(* Logix 5000 project; controller PLC_MCC1201_220AP1 vendor 1 type 14 code 164 rev 35.11; software revision 35.00; part 12 of 25 *)
(* tags used below, declared in another part *)
   B180 : DINT[10];
   BT181_009 : MESSAGE;
   BT181_010 : MESSAGE;
   C183 : COUNTER[3];
   N124 : DINT[414];
   N125 : DINT[414];
   N126 : DINT[103];
   N127 : DINT[997];
   N128 : DINT[997];
   N177_0 : ALIAS FOR N177[0];
   N184 : DINT[50];
   N184_1 : ALIAS FOR N184[1];
   N184_11 : ALIAS FOR N184[11];
   N184_12 : ALIAS FOR N184[12];
   N184_14 : ALIAS FOR N184[14];
   N184_16 : ALIAS FOR N184[16];
   N184_2 : ALIAS FOR N184[2];
   N184_21 : ALIAS FOR N184[21];
   N184_22 : ALIAS FOR N184[22];
   N184_24 : ALIAS FOR N184[24];
   N184_25 : ALIAS FOR N184[25];
   N184_26 : ALIAS FOR N184[26];
   N184_31 : ALIAS FOR N184[31];
   N184_32 : ALIAS FOR N184[32];
   N184_34 : ALIAS FOR N184[34];
   N184_36 : ALIAS FOR N184[36];
   N184_4 : ALIAS FOR N184[4];
   N184_5 : ALIAS FOR N184[5];
   N184_6 : ALIAS FOR N184[6];
   N26 : DINT[1000];
   T182 : TIMER[11];
   TMP_xAlwaysOFF : BOOL;
(* MainProgram, continued *)

ROUTINE _103_LADDER   (* ladder *)
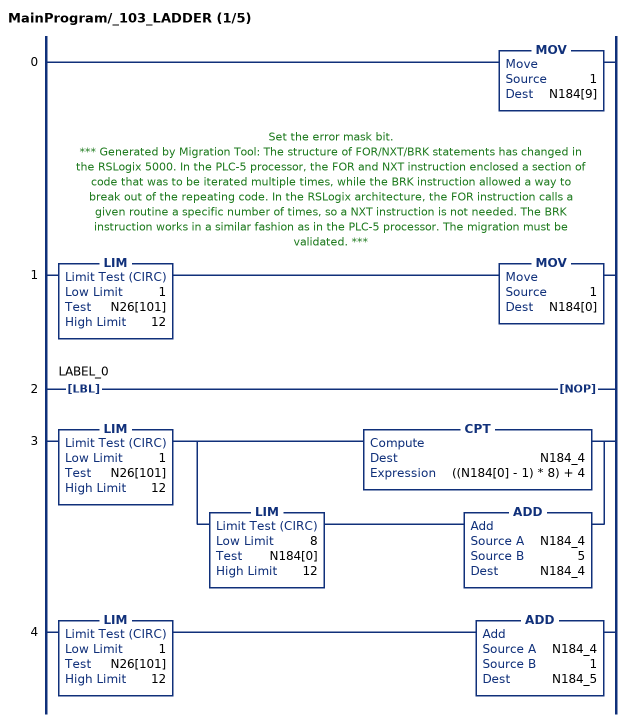
   0: MOV(1,N184[9]);
   // Set the error mask bit.
   // *** Generated by Migration Tool: The structure of FOR/NXT/BRK statements has changed in the RSLogix 5000. In the PLC-5 processor, the FOR and NXT instruction enclosed a section of code that was to be iterated multiple times, while the BRK instruction allowed a way to break out of the repeating code. In the RSLogix architecture, the FOR instruction calls a given routine a specific number of times, so a NXT instruction is not needed. The BRK instruction works in a similar fashion as in the PLC-5 processor. The migration must be validated. ***
   1: LIM(1,N26[101],12)MOV(1,N184[0]);
   2: LBL(LABEL_0)NOP();
   3: LIM(1,N26[101],12)[CPT(N184_4,((N184[0] - 1) * 8) + 4) ,LIM(8,N184[0],12) ADD(N184_4,5,N184_4) ];
   4: LIM(1,N26[101],12)ADD(N184_4,1,N184_5);
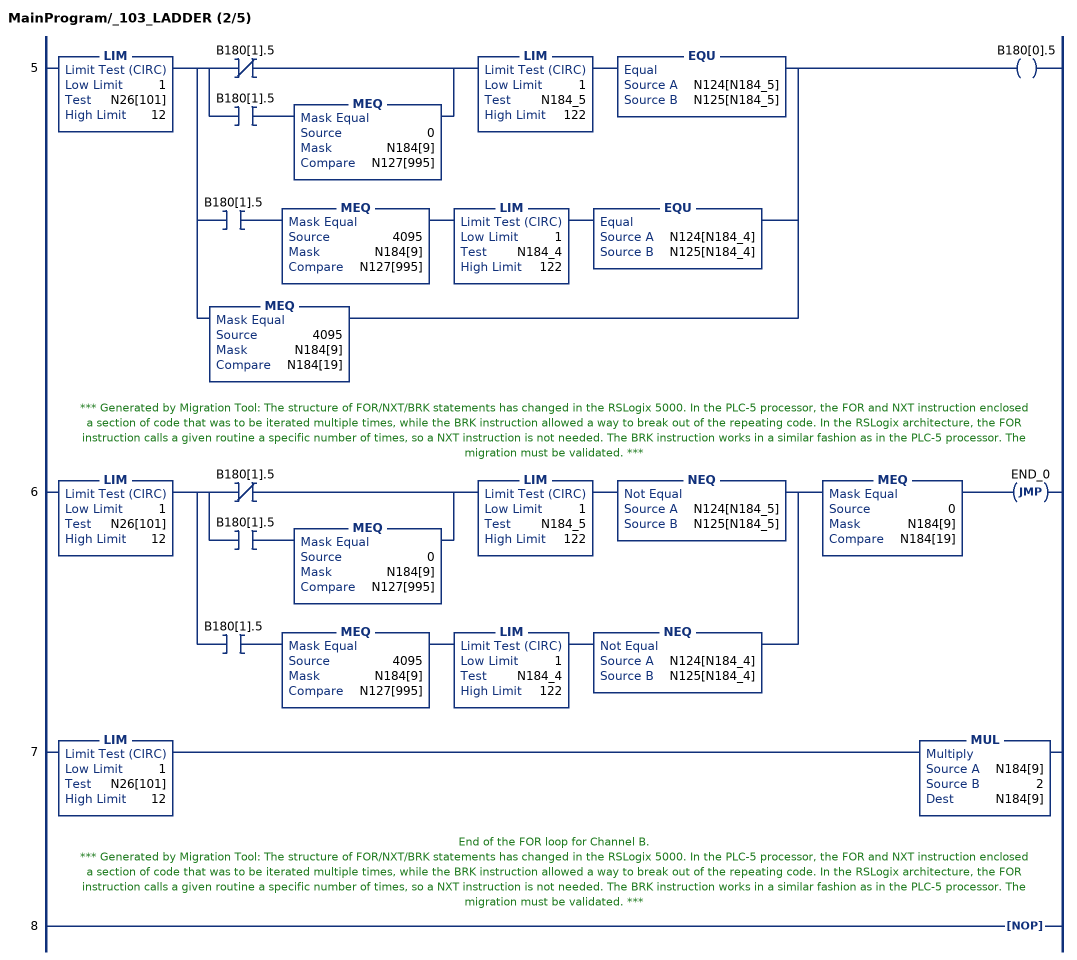
   5: LIM(1,N26[101],12)[[XIO(B180[1].5) ,XIC(B180[1].5) MEQ(0,N184[9],N127[995]) ] LIM(1,N184_5,122) EQU(N124[N184_5],N125[N184_5]) ,XIC(B180[1].5) MEQ(4095,N184[9],N127[995]) LIM(1,N184_4,122) EQU(N124[N184_4],N125[N184_4]) ,MEQ(4095,N184[9],N184[19]) ]OTE(B180[0].5);
   // *** Generated by Migration Tool: The structure of FOR/NXT/BRK statements has changed in the RSLogix 5000. In the PLC-5 processor, the FOR and NXT instruction enclosed a section of code that was to be iterated multiple times, while the BRK instruction allowed a way to break out of the repeating code. In the RSLogix architecture, the FOR instruction calls a given routine a specific number of times, so a NXT instruction is not needed. The BRK instruction works in a similar fashion as in the PLC-5 processor. The migration must be validated. ***
   6: LIM(1,N26[101],12)[[XIO(B180[1].5) ,XIC(B180[1].5) MEQ(0,N184[9],N127[995]) ] LIM(1,N184_5,122) NEQ(N124[N184_5],N125[N184_5]) ,XIC(B180[1].5) MEQ(4095,N184[9],N127[995]) LIM(1,N184_4,122) NEQ(N124[N184_4],N125[N184_4]) ]MEQ(0,N184[9],N184[19])JMP(END_0);
   7: LIM(1,N26[101],12)MUL(N184[9],2,N184[9]);
   // End of the FOR loop for Channel B.
   // *** Generated by Migration Tool: The structure of FOR/NXT/BRK statements has changed in the RSLogix 5000. In the PLC-5 processor, the FOR and NXT instruction enclosed a section of code that was to be iterated multiple times, while the BRK instruction allowed a way to break out of the repeating code. In the RSLogix architecture, the FOR instruction calls a given routine a specific number of times, so a NXT instruction is not needed. The BRK instruction works in a similar fashion as in the PLC-5 processor. The migration must be validated. ***
   8: NOP();
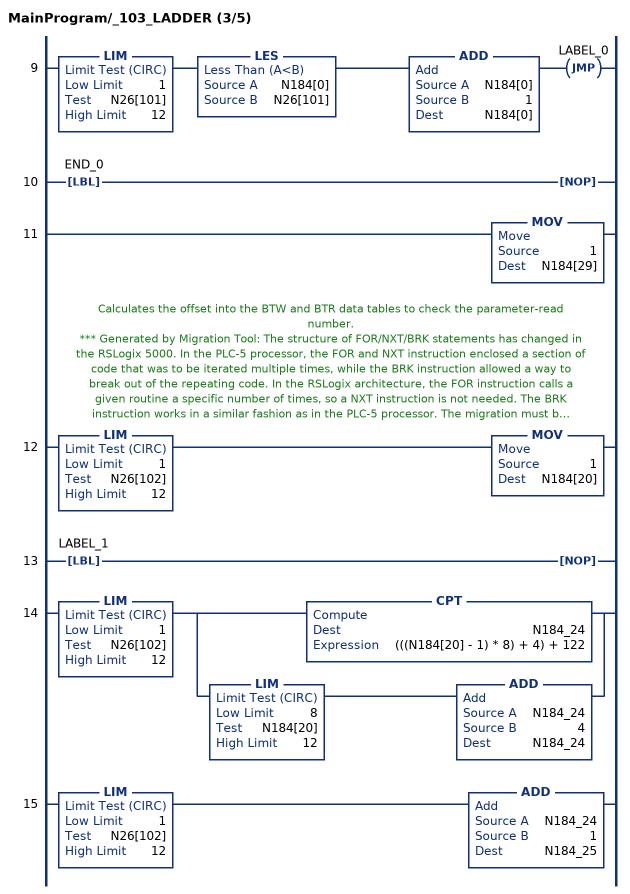
   9: LIM(1,N26[101],12)LES(N184[0],N26[101])ADD(N184[0],1,N184[0])JMP(LABEL_0);
   10: LBL(END_0)NOP();
   11: MOV(1,N184[29]);
   // Calculates the offset into the BTW and BTR data tables to check the parameter-read number.
   // *** Generated by Migration Tool: The structure of FOR/NXT/BRK statements has changed in the RSLogix 5000. In the PLC-5 processor, the FOR and NXT instruction enclosed a section of code that was to be iterated multiple times, while the BRK instruction allowed a way to break out of the repeating code. In the RSLogix architecture, the FOR instruction calls a given routine a specific number of times, so a NXT instruction is not needed. The BRK instruction works in a similar fashion as in the PLC-5 processor. The migration must be validated. ***
   12: LIM(1,N26[102],12)MOV(1,N184[20]);
   13: LBL(LABEL_1)NOP();
   14: LIM(1,N26[102],12)[CPT(N184_24,(((N184[20] - 1) * 8) + 4) + 122) ,LIM(8,N184[20],12) ADD(N184_24,4,N184_24) ];
   15: LIM(1,N26[102],12)ADD(N184_24,1,N184_25);
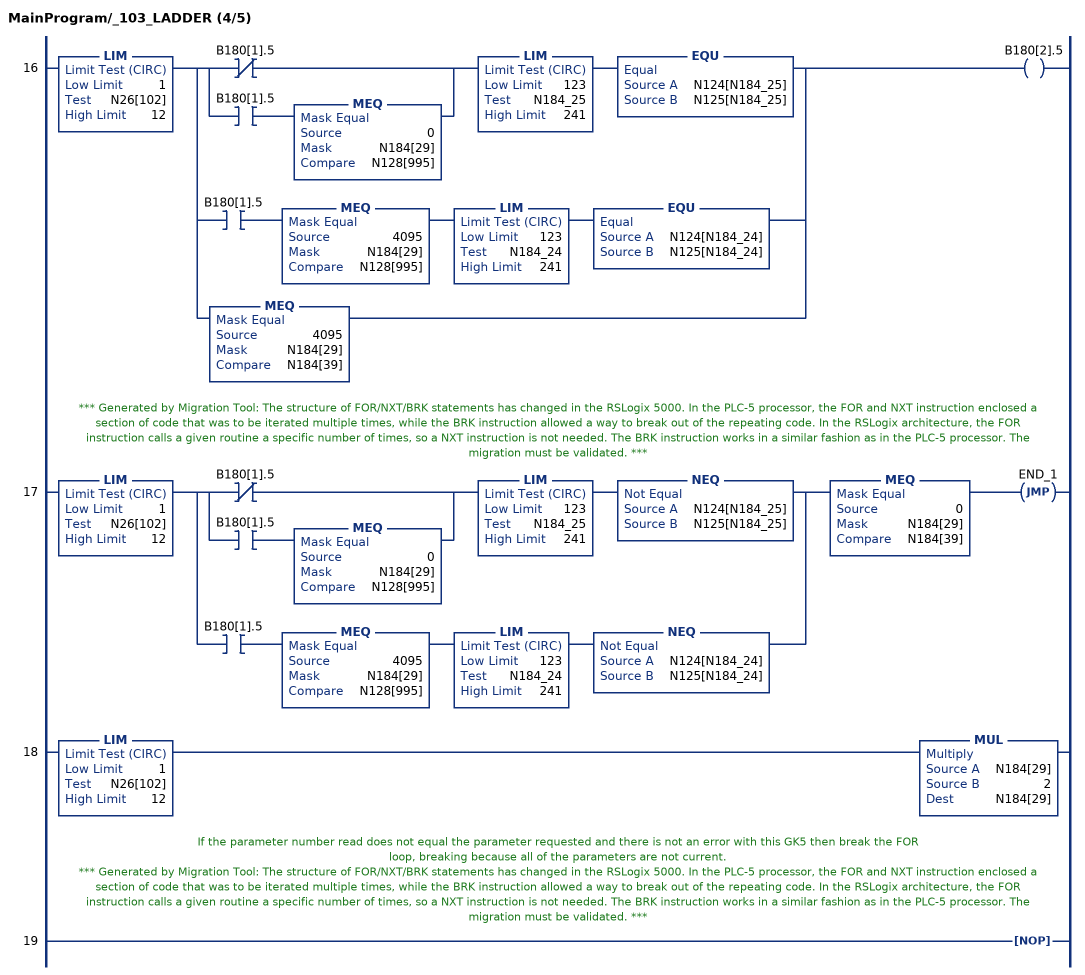
   16: LIM(1,N26[102],12)[[XIO(B180[1].5) ,XIC(B180[1].5) MEQ(0,N184[29],N128[995]) ] LIM(123,N184_25,241) EQU(N124[N184_25],N125[N184_25]) ,XIC(B180[1].5) MEQ(4095,N184[29],N128[995]) LIM(123,N184_24,241) EQU(N124[N184_24],N125[N184_24]) ,MEQ(4095,N184[29],N184[39]) ]OTE(B180[2].5);
   // *** Generated by Migration Tool: The structure of FOR/NXT/BRK statements has changed in the RSLogix 5000. In the PLC-5 processor, the FOR and NXT instruction enclosed a section of code that was to be iterated multiple times, while the BRK instruction allowed a way to break out of the repeating code. In the RSLogix architecture, the FOR instruction calls a given routine a specific number of times, so a NXT instruction is not needed. The BRK instruction works in a similar fashion as in the PLC-5 processor. The migration must be validated. ***
   17: LIM(1,N26[102],12)[[XIO(B180[1].5) ,XIC(B180[1].5) MEQ(0,N184[29],N128[995]) ] LIM(123,N184_25,241) NEQ(N124[N184_25],N125[N184_25]) ,XIC(B180[1].5) MEQ(4095,N184[29],N128[995]) LIM(123,N184_24,241) NEQ(N124[N184_24],N125[N184_24]) ]MEQ(0,N184[29],N184[39])JMP(END_1);
   18: LIM(1,N26[102],12)MUL(N184[29],2,N184[29]);
   // If the parameter number read does not equal the parameter requested and there is not an error with this GK5 then break the FOR
   // loop, breaking because all of the parameters are not current.
   // *** Generated by Migration Tool: The structure of FOR/NXT/BRK statements has changed in the RSLogix 5000. In the PLC-5 processor, the FOR and NXT instruction enclosed a section of code that was to be iterated multiple times, while the BRK instruction allowed a way to break out of the repeating code. In the RSLogix architecture, the FOR instruction calls a given routine a specific number of times, so a NXT instruction is not needed. The BRK instruction works in a similar fashion as in the PLC-5 processor. The migration must be validated. ***
   19: NOP();
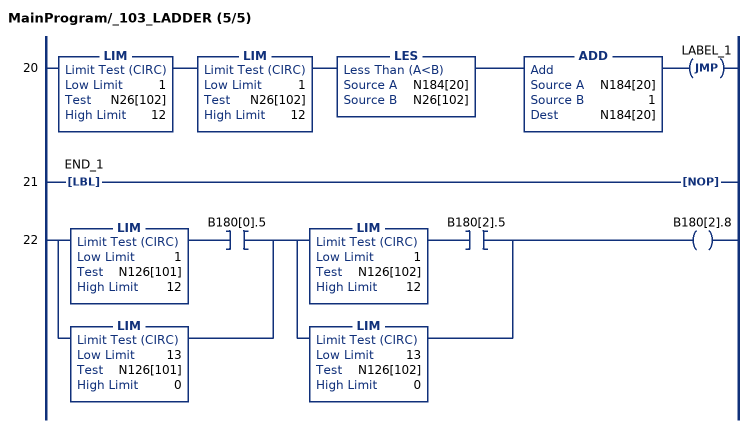
   20: LIM(1,N26[102],12)LIM(1,N26[102],12)LES(N184[20],N26[102])ADD(N184[20],1,N184[20])JMP(LABEL_1);
   21: LBL(END_1)NOP();
   22: [LIM(1,N126[101],12) XIC(B180[0].5) ,LIM(13,N126[101],0) ][LIM(1,N126[102],12) XIC(B180[2].5) ,LIM(13,N126[102],0) ]OTE(B180[2].8);
END_ROUTINE

ROUTINE _104_LADDER   (* ladder *)
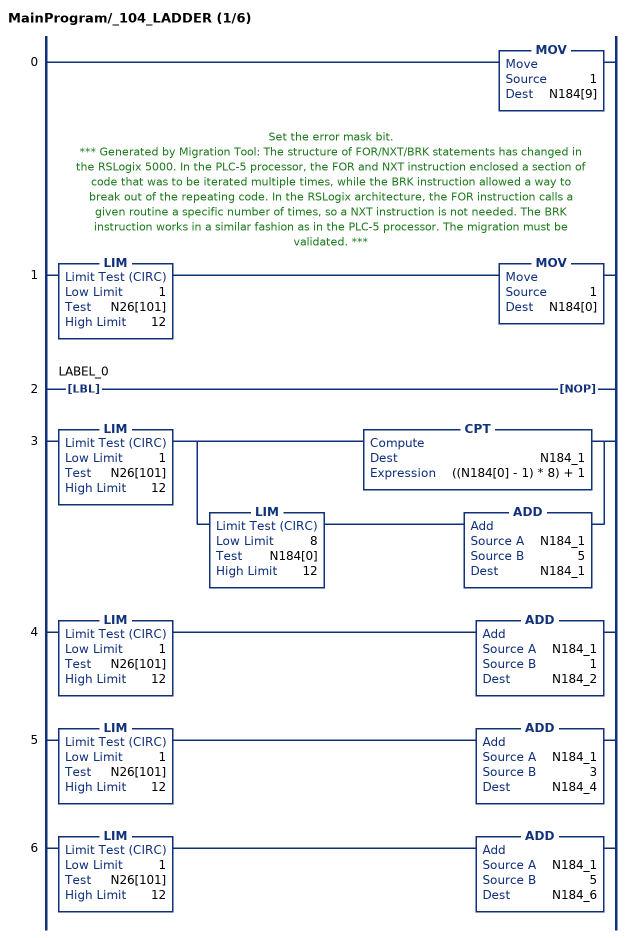
   0: MOV(1,N184[9]);
   // Set the error mask bit.
   // *** Generated by Migration Tool: The structure of FOR/NXT/BRK statements has changed in the RSLogix 5000. In the PLC-5 processor, the FOR and NXT instruction enclosed a section of code that was to be iterated multiple times, while the BRK instruction allowed a way to break out of the repeating code. In the RSLogix architecture, the FOR instruction calls a given routine a specific number of times, so a NXT instruction is not needed. The BRK instruction works in a similar fashion as in the PLC-5 processor. The migration must be validated. ***
   1: LIM(1,N26[101],12)MOV(1,N184[0]);
   2: LBL(LABEL_0)NOP();
   3: LIM(1,N26[101],12)[CPT(N184_1,((N184[0] - 1) * 8) + 1) ,LIM(8,N184[0],12) ADD(N184_1,5,N184_1) ];
   4: LIM(1,N26[101],12)ADD(N184_1,1,N184_2);
   5: LIM(1,N26[101],12)ADD(N184_1,3,N184_4);
   6: LIM(1,N26[101],12)ADD(N184_1,5,N184_6);
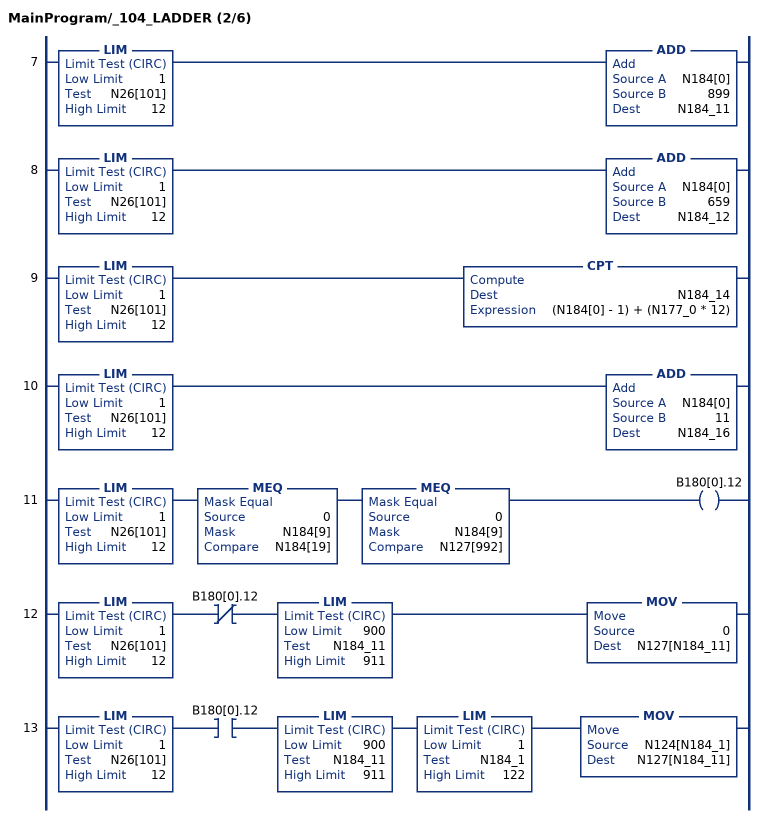
   7: LIM(1,N26[101],12)ADD(N184[0],899,N184_11);
   8: LIM(1,N26[101],12)ADD(N184[0],659,N184_12);
   9: LIM(1,N26[101],12)CPT(N184_14,(N184[0] - 1) + (N177_0 * 12));
   10: LIM(1,N26[101],12)ADD(N184[0],11,N184_16);
   11: LIM(1,N26[101],12)MEQ(0,N184[9],N184[19])MEQ(0,N184[9],N127[992])OTE(B180[0].12);
   12: LIM(1,N26[101],12)XIO(B180[0].12)LIM(900,N184_11,911)MOV(0,N127[N184_11]);
   13: LIM(1,N26[101],12)XIC(B180[0].12)LIM(900,N184_11,911)LIM(1,N184_1,122)MOV(N124[N184_1],N127[N184_11]);
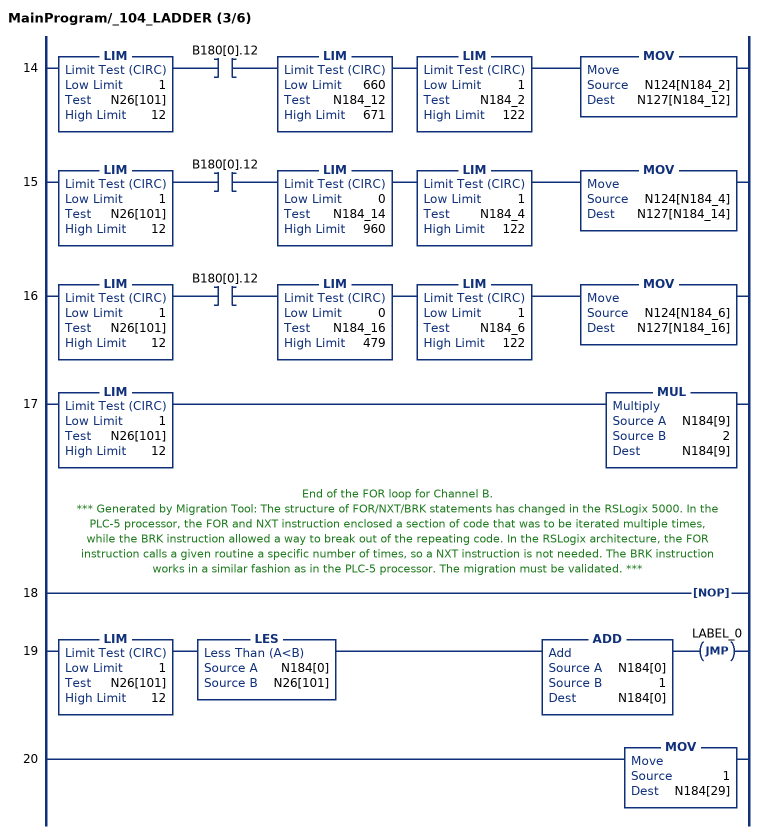
   14: LIM(1,N26[101],12)XIC(B180[0].12)LIM(660,N184_12,671)LIM(1,N184_2,122)MOV(N124[N184_2],N127[N184_12]);
   15: LIM(1,N26[101],12)XIC(B180[0].12)LIM(0,N184_14,960)LIM(1,N184_4,122)MOV(N124[N184_4],N127[N184_14]);
   16: LIM(1,N26[101],12)XIC(B180[0].12)LIM(0,N184_16,479)LIM(1,N184_6,122)MOV(N124[N184_6],N127[N184_16]);
   17: LIM(1,N26[101],12)MUL(N184[9],2,N184[9]);
   // End of the FOR loop for Channel B.
   // *** Generated by Migration Tool: The structure of FOR/NXT/BRK statements has changed in the RSLogix 5000. In the PLC-5 processor, the FOR and NXT instruction enclosed a section of code that was to be iterated multiple times, while the BRK instruction allowed a way to break out of the repeating code. In the RSLogix architecture, the FOR instruction calls a given routine a specific number of times, so a NXT instruction is not needed. The BRK instruction works in a similar fashion as in the PLC-5 processor. The migration must be validated. ***
   18: NOP();
   19: LIM(1,N26[101],12)LES(N184[0],N26[101])ADD(N184[0],1,N184[0])JMP(LABEL_0);
   20: MOV(1,N184[29]);
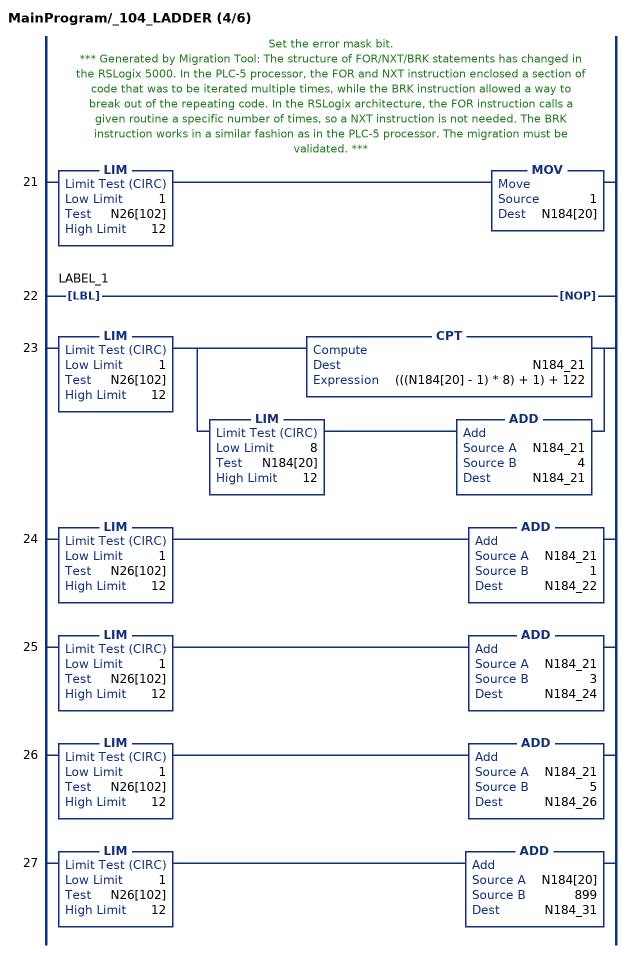
   // Set the error mask bit.
   // *** Generated by Migration Tool: The structure of FOR/NXT/BRK statements has changed in the RSLogix 5000. In the PLC-5 processor, the FOR and NXT instruction enclosed a section of code that was to be iterated multiple times, while the BRK instruction allowed a way to break out of the repeating code. In the RSLogix architecture, the FOR instruction calls a given routine a specific number of times, so a NXT instruction is not needed. The BRK instruction works in a similar fashion as in the PLC-5 processor. The migration must be validated. ***
   21: LIM(1,N26[102],12)MOV(1,N184[20]);
   22: LBL(LABEL_1)NOP();
   23: LIM(1,N26[102],12)[CPT(N184_21,(((N184[20] - 1) * 8) + 1) + 122) ,LIM(8,N184[20],12) ADD(N184_21,4,N184_21) ];
   24: LIM(1,N26[102],12)ADD(N184_21,1,N184_22);
   25: LIM(1,N26[102],12)ADD(N184_21,3,N184_24);
   26: LIM(1,N26[102],12)ADD(N184_21,5,N184_26);
   27: LIM(1,N26[102],12)ADD(N184[20],899,N184_31);
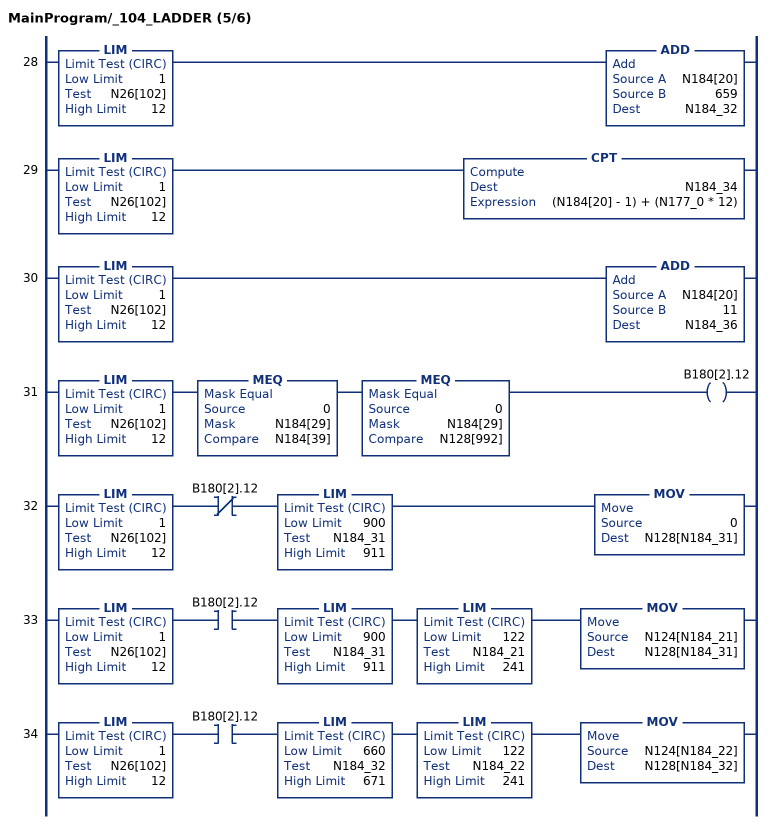
   28: LIM(1,N26[102],12)ADD(N184[20],659,N184_32);
   29: LIM(1,N26[102],12)CPT(N184_34,(N184[20] - 1) + (N177_0 * 12));
   30: LIM(1,N26[102],12)ADD(N184[20],11,N184_36);
   31: LIM(1,N26[102],12)MEQ(0,N184[29],N184[39])MEQ(0,N184[29],N128[992])OTE(B180[2].12);
   32: LIM(1,N26[102],12)XIO(B180[2].12)LIM(900,N184_31,911)MOV(0,N128[N184_31]);
   33: LIM(1,N26[102],12)XIC(B180[2].12)LIM(900,N184_31,911)LIM(122,N184_21,241)MOV(N124[N184_21],N128[N184_31]);
   34: LIM(1,N26[102],12)XIC(B180[2].12)LIM(660,N184_32,671)LIM(122,N184_22,241)MOV(N124[N184_22],N128[N184_32]);
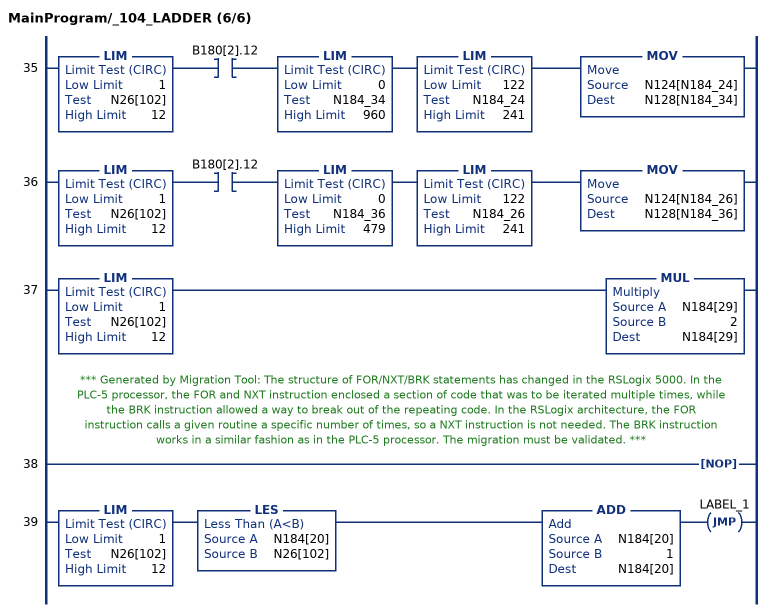
   35: LIM(1,N26[102],12)XIC(B180[2].12)LIM(0,N184_34,960)LIM(122,N184_24,241)MOV(N124[N184_24],N128[N184_34]);
   36: LIM(1,N26[102],12)XIC(B180[2].12)LIM(0,N184_36,479)LIM(122,N184_26,241)MOV(N124[N184_26],N128[N184_36]);
   37: LIM(1,N26[102],12)MUL(N184[29],2,N184[29]);
   // *** Generated by Migration Tool: The structure of FOR/NXT/BRK statements has changed in the RSLogix 5000. In the PLC-5 processor, the FOR and NXT instruction enclosed a section of code that was to be iterated multiple times, while the BRK instruction allowed a way to break out of the repeating code. In the RSLogix architecture, the FOR instruction calls a given routine a specific number of times, so a NXT instruction is not needed. The BRK instruction works in a similar fashion as in the PLC-5 processor. The migration must be validated. ***
   38: NOP();
   39: LIM(1,N26[102],12)LES(N184[20],N26[102])ADD(N184[20],1,N184[20])JMP(LABEL_1);
END_ROUTINE

ROUTINE _105_LADDER   (* ladder *)
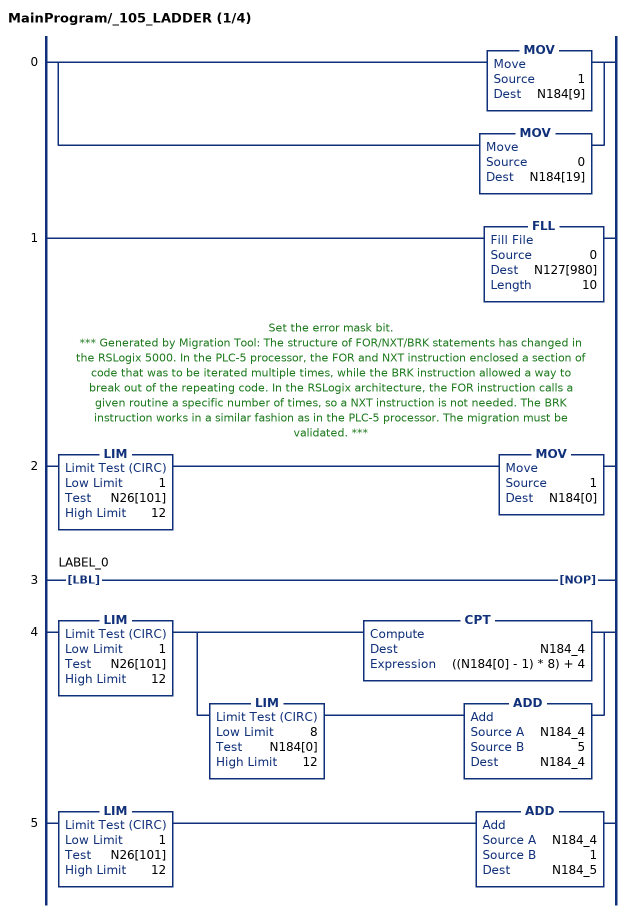
   0: [MOV(1,N184[9]) ,MOV(0,N184[19]) ];
   1: FLL(0,N127[980],10);
   // Set the error mask bit.
   // *** Generated by Migration Tool: The structure of FOR/NXT/BRK statements has changed in the RSLogix 5000. In the PLC-5 processor, the FOR and NXT instruction enclosed a section of code that was to be iterated multiple times, while the BRK instruction allowed a way to break out of the repeating code. In the RSLogix architecture, the FOR instruction calls a given routine a specific number of times, so a NXT instruction is not needed. The BRK instruction works in a similar fashion as in the PLC-5 processor. The migration must be validated. ***
   2: LIM(1,N26[101],12)MOV(1,N184[0]);
   3: LBL(LABEL_0)NOP();
   4: LIM(1,N26[101],12)[CPT(N184_4,((N184[0] - 1) * 8) + 4) ,LIM(8,N184[0],12) ADD(N184_4,5,N184_4) ];
   5: LIM(1,N26[101],12)ADD(N184_4,1,N184_5);
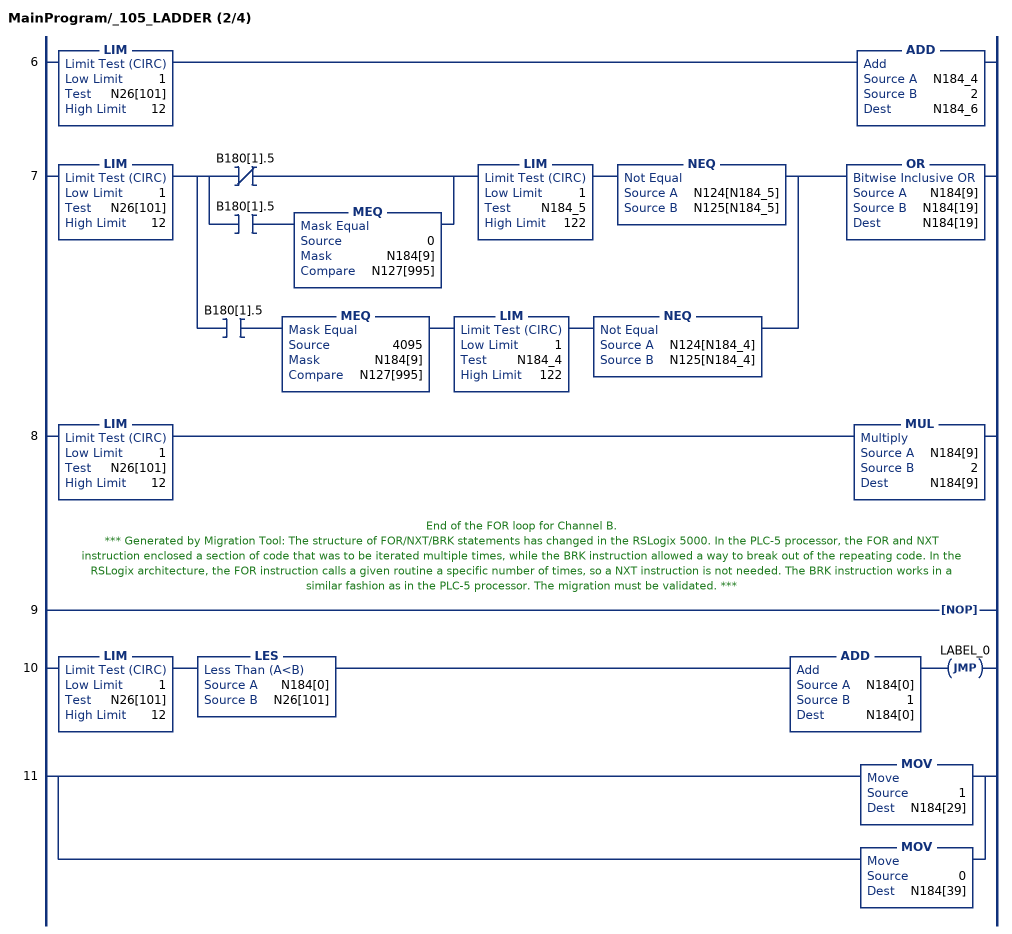
   6: LIM(1,N26[101],12)ADD(N184_4,2,N184_6);
   7: LIM(1,N26[101],12)[[XIO(B180[1].5) ,XIC(B180[1].5) MEQ(0,N184[9],N127[995]) ] LIM(1,N184_5,122) NEQ(N124[N184_5],N125[N184_5]) ,XIC(B180[1].5) MEQ(4095,N184[9],N127[995]) LIM(1,N184_4,122) NEQ(N124[N184_4],N125[N184_4]) ]OR(N184[9],N184[19],N184[19]);
   8: LIM(1,N26[101],12)MUL(N184[9],2,N184[9]);
   // End of the FOR loop for Channel B.
   // *** Generated by Migration Tool: The structure of FOR/NXT/BRK statements has changed in the RSLogix 5000. In the PLC-5 processor, the FOR and NXT instruction enclosed a section of code that was to be iterated multiple times, while the BRK instruction allowed a way to break out of the repeating code. In the RSLogix architecture, the FOR instruction calls a given routine a specific number of times, so a NXT instruction is not needed. The BRK instruction works in a similar fashion as in the PLC-5 processor. The migration must be validated. ***
   9: NOP();
   10: LIM(1,N26[101],12)LES(N184[0],N26[101])ADD(N184[0],1,N184[0])JMP(LABEL_0);
   11: [MOV(1,N184[29]) ,MOV(0,N184[39]) ];
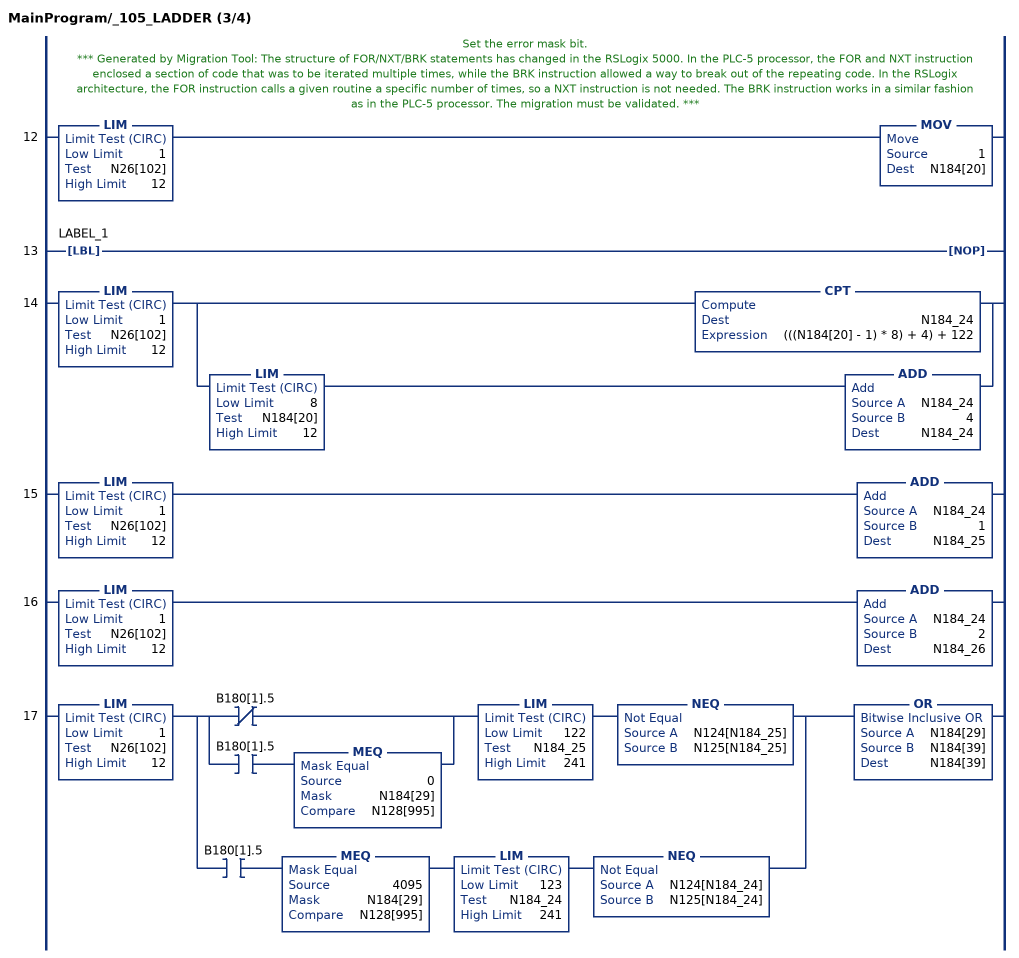
   // Set the error mask bit.
   // *** Generated by Migration Tool: The structure of FOR/NXT/BRK statements has changed in the RSLogix 5000. In the PLC-5 processor, the FOR and NXT instruction enclosed a section of code that was to be iterated multiple times, while the BRK instruction allowed a way to break out of the repeating code. In the RSLogix architecture, the FOR instruction calls a given routine a specific number of times, so a NXT instruction is not needed. The BRK instruction works in a similar fashion as in the PLC-5 processor. The migration must be validated. ***
   12: LIM(1,N26[102],12)MOV(1,N184[20]);
   13: LBL(LABEL_1)NOP();
   14: LIM(1,N26[102],12)[CPT(N184_24,(((N184[20] - 1) * 8) + 4) + 122) ,LIM(8,N184[20],12) ADD(N184_24,4,N184_24) ];
   15: LIM(1,N26[102],12)ADD(N184_24,1,N184_25);
   16: LIM(1,N26[102],12)ADD(N184_24,2,N184_26);
   17: LIM(1,N26[102],12)[[XIO(B180[1].5) ,XIC(B180[1].5) MEQ(0,N184[29],N128[995]) ] LIM(122,N184_25,241) NEQ(N124[N184_25],N125[N184_25]) ,XIC(B180[1].5) MEQ(4095,N184[29],N128[995]) LIM(123,N184_24,241) NEQ(N124[N184_24],N125[N184_24]) ]OR(N184[29],N184[39],N184[39]);
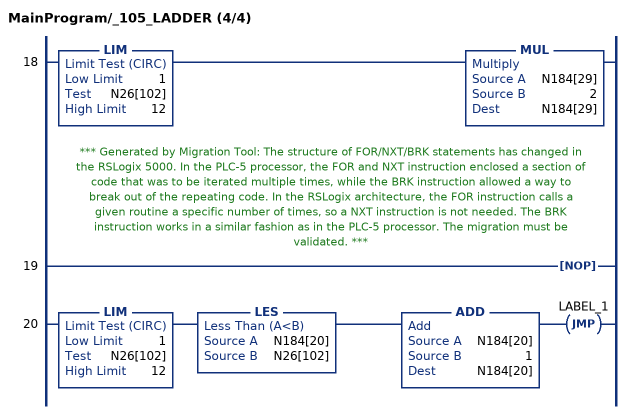
   18: LIM(1,N26[102],12)MUL(N184[29],2,N184[29]);
   // *** Generated by Migration Tool: The structure of FOR/NXT/BRK statements has changed in the RSLogix 5000. In the PLC-5 processor, the FOR and NXT instruction enclosed a section of code that was to be iterated multiple times, while the BRK instruction allowed a way to break out of the repeating code. In the RSLogix architecture, the FOR instruction calls a given routine a specific number of times, so a NXT instruction is not needed. The BRK instruction works in a similar fashion as in the PLC-5 processor. The migration must be validated. ***
   19: NOP();
   20: LIM(1,N26[102],12)LES(N184[20],N26[102])ADD(N184[20],1,N184[20])JMP(LABEL_1);
END_ROUTINE

ROUTINE _106_LADDER   (* ladder *)
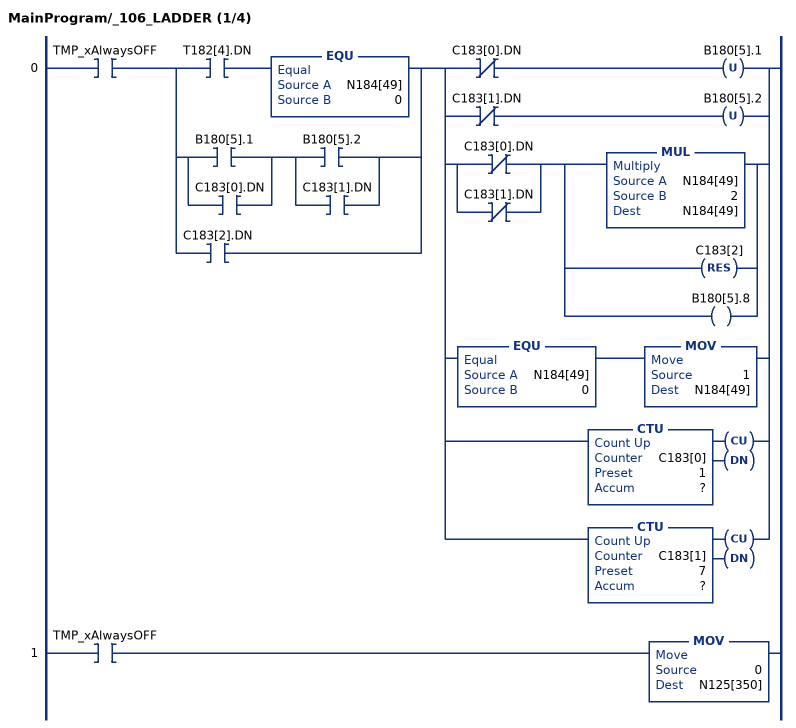
   0: XIC(TMP_xAlwaysOFF)[XIC(T182[4].DN) EQU(N184[49],0) ,[XIC(B180[5].1) ,XIC(C183[0].DN) ] [XIC(B180[5].2) ,XIC(C183[1].DN) ] ,XIC(C183[2].DN) ][XIO(C183[0].DN) OTU(B180[5].1) ,XIO(C183[1].DN) OTU(B180[5].2) ,[XIO(C183[0].DN) ,XIO(C183[1].DN) ] [MUL(N184[49],2,N184[49]) ,RES(C183[2]) ,OTE(B180[5].8) ] ,EQU(N184[49],0) MOV(1,N184[49]) ,CTU(C183[0],?,?) ,CTU(C183[1],?,?) ];
   1: XIC(TMP_xAlwaysOFF)MOV(0,N125[350]);
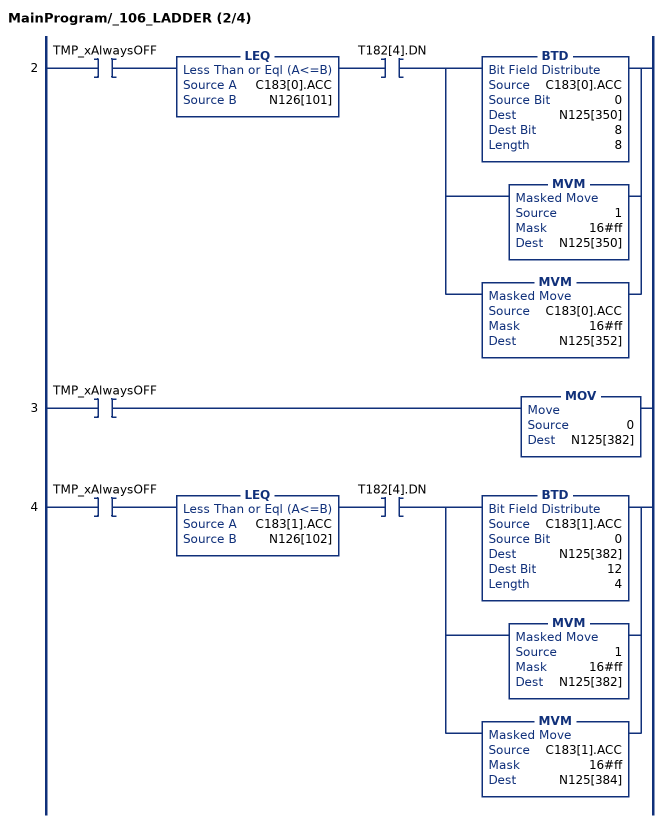
   2: XIC(TMP_xAlwaysOFF)LEQ(C183[0].ACC,N126[101])XIC(T182[4].DN)[BTD(C183[0].ACC,0,N125[350],8,8) ,MVM(1,16#ff,N125[350]) ,MVM(C183[0].ACC,16#ff,N125[352]) ];
   3: XIC(TMP_xAlwaysOFF)MOV(0,N125[382]);
   4: XIC(TMP_xAlwaysOFF)LEQ(C183[1].ACC,N126[102])XIC(T182[4].DN)[BTD(C183[1].ACC,0,N125[382],12,4) ,MVM(1,16#ff,N125[382]) ,MVM(C183[1].ACC,16#ff,N125[384]) ];
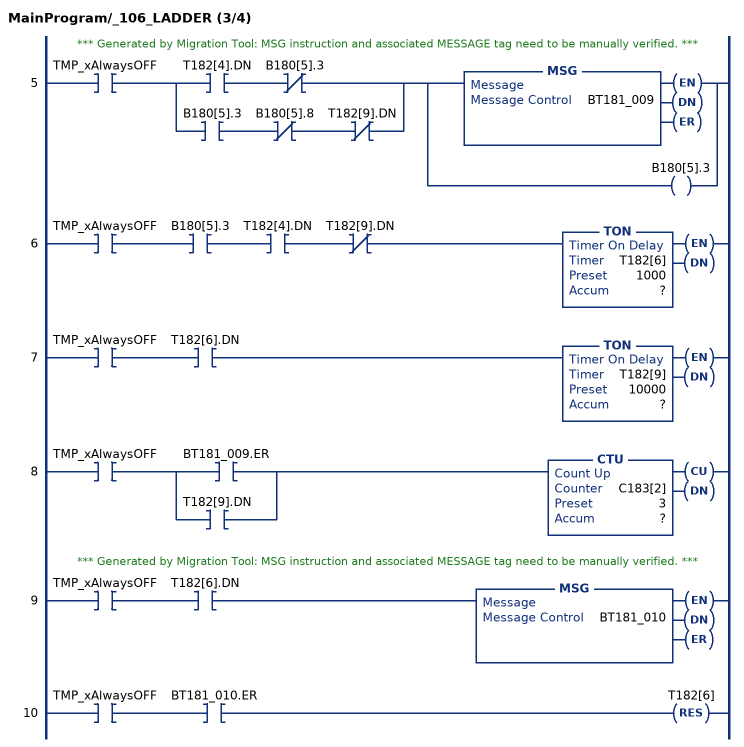
   // *** Generated by Migration Tool: MSG instruction and associated MESSAGE tag need to be manually verified. ***
   5: XIC(TMP_xAlwaysOFF)[XIC(T182[4].DN) XIO(B180[5].3) ,XIC(B180[5].3) XIO(B180[5].8) XIO(T182[9].DN) ][MSG(BT181_009) ,OTE(B180[5].3) ];
   6: XIC(TMP_xAlwaysOFF)XIC(B180[5].3)XIC(T182[4].DN)XIO(T182[9].DN)TON(T182[6],?,?);
   7: XIC(TMP_xAlwaysOFF)XIC(T182[6].DN)TON(T182[9],?,?);
   8: XIC(TMP_xAlwaysOFF)[XIC(BT181_009.ER) ,XIC(T182[9].DN) ]CTU(C183[2],?,?);
   // *** Generated by Migration Tool: MSG instruction and associated MESSAGE tag need to be manually verified. ***
   9: XIC(TMP_xAlwaysOFF)XIC(T182[6].DN)MSG(BT181_010);
   10: XIC(TMP_xAlwaysOFF)XIC(BT181_010.ER)RES(T182[6]);
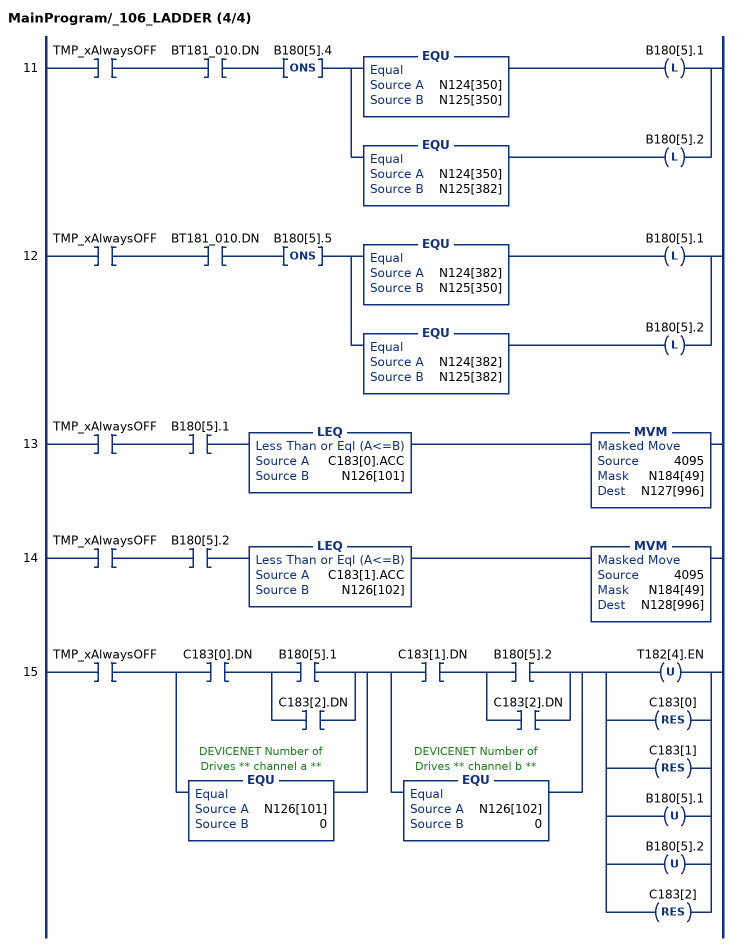
   11: XIC(TMP_xAlwaysOFF)XIC(BT181_010.DN)ONS(B180[5].4)[EQU(N124[350],N125[350]) OTL(B180[5].1) ,EQU(N124[350],N125[382]) OTL(B180[5].2) ];
   12: XIC(TMP_xAlwaysOFF)XIC(BT181_010.DN)ONS(B180[5].5)[EQU(N124[382],N125[350]) OTL(B180[5].1) ,EQU(N124[382],N125[382]) OTL(B180[5].2) ];
   13: XIC(TMP_xAlwaysOFF)XIC(B180[5].1)LEQ(C183[0].ACC,N126[101])MVM(4095,N184[49],N127[996]);
   14: XIC(TMP_xAlwaysOFF)XIC(B180[5].2)LEQ(C183[1].ACC,N126[102])MVM(4095,N184[49],N128[996]);
   15: XIC(TMP_xAlwaysOFF)[XIC(C183[0].DN) [XIC(B180[5].1) ,XIC(C183[2].DN) ] ,EQU(N126[101],0) ][XIC(C183[1].DN) [XIC(B180[5].2) ,XIC(C183[2].DN) ] ,EQU(N126[102],0) ][OTU(T182[4].EN) ,RES(C183[0]) ,RES(C183[1]) ,OTU(B180[5].1) ,OTU(B180[5].2) ,RES(C183[2]) ];
END_ROUTINE
